REGION Network 297: CARRIER POWER UNIT DC LINK UNDERVOLTAGE
   RUNG wire#powerrail
      { S7_Templates := "SrcType := Word" } EQ_Contact(in1 := "DB101_DB_SDC_FAULTS".Carrier_Fault[8], in2 := 182)
      Coil( "DB302_HMI_Faults".Carrier8_Faults_1.%X11 )
   END_RUNG
   // the same network as SCL:
   "DB302_HMI_Faults".Carrier8_Faults_1.%X11 := "DB101_DB_SDC_FAULTS".Carrier_Fault[8] = 182;
END_REGION

REGION Network 298: CARRIER POWER UNIT LINE PHASE FAILURE
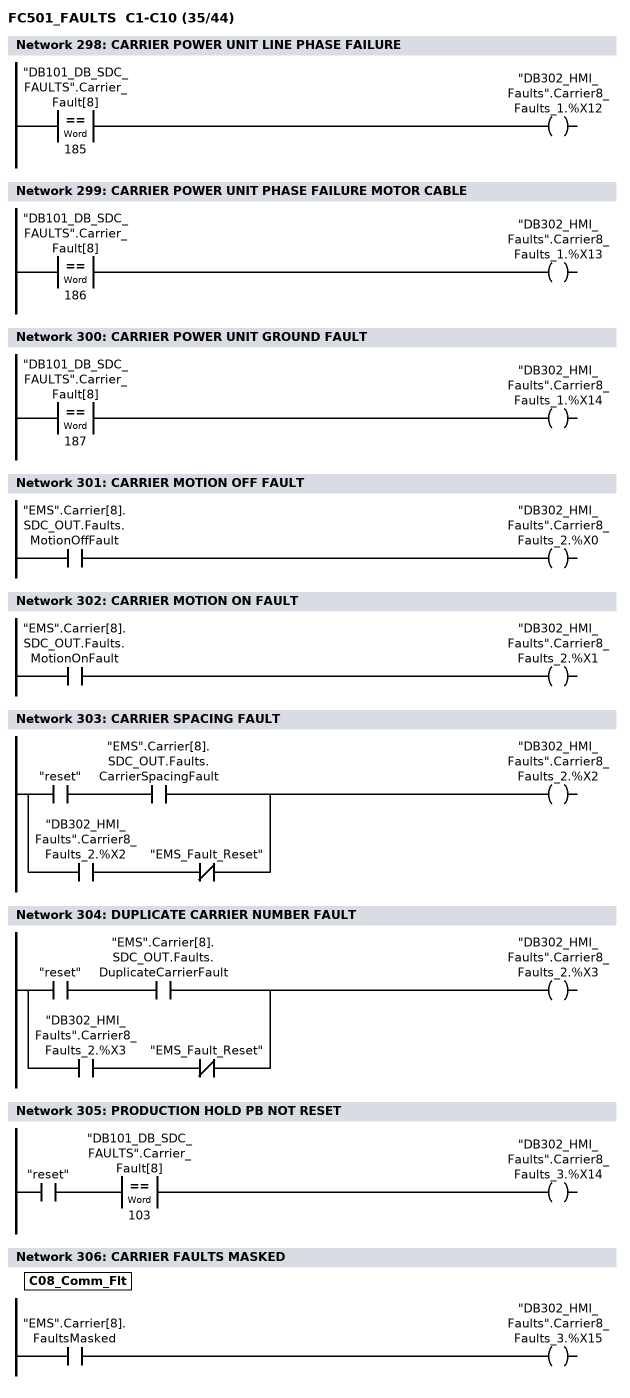
   RUNG wire#powerrail
      { S7_Templates := "SrcType := Word" } EQ_Contact(in1 := "DB101_DB_SDC_FAULTS".Carrier_Fault[8], in2 := 185)
      Coil( "DB302_HMI_Faults".Carrier8_Faults_1.%X12 )
   END_RUNG
   // the same network as SCL:
   "DB302_HMI_Faults".Carrier8_Faults_1.%X12 := "DB101_DB_SDC_FAULTS".Carrier_Fault[8] = 185;
END_REGION

REGION Network 299: CARRIER POWER UNIT PHASE FAILURE MOTOR CABLE
   RUNG wire#powerrail
      { S7_Templates := "SrcType := Word" } EQ_Contact(in1 := "DB101_DB_SDC_FAULTS".Carrier_Fault[8], in2 := 186)
      Coil( "DB302_HMI_Faults".Carrier8_Faults_1.%X13 )
   END_RUNG
   // the same network as SCL:
   "DB302_HMI_Faults".Carrier8_Faults_1.%X13 := "DB101_DB_SDC_FAULTS".Carrier_Fault[8] = 186;
END_REGION

REGION Network 300: CARRIER POWER UNIT GROUND FAULT
   RUNG wire#powerrail
      { S7_Templates := "SrcType := Word" } EQ_Contact(in1 := "DB101_DB_SDC_FAULTS".Carrier_Fault[8], in2 := 187)
      Coil( "DB302_HMI_Faults".Carrier8_Faults_1.%X14 )
   END_RUNG
   // the same network as SCL:
   "DB302_HMI_Faults".Carrier8_Faults_1.%X14 := "DB101_DB_SDC_FAULTS".Carrier_Fault[8] = 187;
END_REGION

REGION Network 301: CARRIER MOTION OFF FAULT
   RUNG wire#powerrail
      Contact( "EMS".Carrier[8].SDC_OUT.Faults.MotionOffFault )
      Coil( "DB302_HMI_Faults".Carrier8_Faults_2.%X0 )
   END_RUNG
   // the same network as SCL:
   "DB302_HMI_Faults".Carrier8_Faults_2.%X0 := "EMS".Carrier[8].SDC_OUT.Faults.MotionOffFault;
END_REGION

REGION Network 302: CARRIER MOTION ON FAULT
   RUNG wire#powerrail
      Contact( "EMS".Carrier[8].SDC_OUT.Faults.MotionOnFault )
      Coil( "DB302_HMI_Faults".Carrier8_Faults_2.%X1 )
   END_RUNG
   // the same network as SCL:
   "DB302_HMI_Faults".Carrier8_Faults_2.%X1 := "EMS".Carrier[8].SDC_OUT.Faults.MotionOnFault;
END_REGION

REGION Network 303: CARRIER SPACING FAULT
   RUNG wire#powerrail
      Contact( "reset" )
      Contact( "EMS".Carrier[8].SDC_OUT.Faults.CarrierSpacingFault )
      wire#w1
      Coil( "DB302_HMI_Faults".Carrier8_Faults_2.%X2 )
   END_RUNG
   RUNG wire#powerrail
      Contact( "DB302_HMI_Faults".Carrier8_Faults_2.%X2 )
      I_Contact( "EMS_Fault_Reset" )
   END_RUNG wire#w1
   // the same network as SCL:
   "DB302_HMI_Faults".Carrier8_Faults_2.%X2 := ("reset" AND "EMS".Carrier[8].SDC_OUT.Faults.CarrierSpacingFault) OR ("DB302_HMI_Faults".Carrier8_Faults_2.%X2 AND NOT "EMS_Fault_Reset");
END_REGION

REGION Network 304: DUPLICATE CARRIER NUMBER FAULT
   RUNG wire#powerrail
      Contact( "reset" )
      Contact( "EMS".Carrier[8].SDC_OUT.Faults.DuplicateCarrierFault )
      wire#w1
      Coil( "DB302_HMI_Faults".Carrier8_Faults_2.%X3 )
   END_RUNG
   RUNG wire#powerrail
      Contact( "DB302_HMI_Faults".Carrier8_Faults_2.%X3 )
      I_Contact( "EMS_Fault_Reset" )
   END_RUNG wire#w1
   // the same network as SCL:
   "DB302_HMI_Faults".Carrier8_Faults_2.%X3 := ("reset" AND "EMS".Carrier[8].SDC_OUT.Faults.DuplicateCarrierFault) OR ("DB302_HMI_Faults".Carrier8_Faults_2.%X3 AND NOT "EMS_Fault_Reset");
END_REGION

REGION Network 305: PRODUCTION HOLD PB NOT RESET
   RUNG wire#powerrail
      Contact( "reset" )
      { S7_Templates := "SrcType := Word" } EQ_Contact(in1 := "DB101_DB_SDC_FAULTS".Carrier_Fault[8], in2 := 103)
      Coil( "DB302_HMI_Faults".Carrier8_Faults_3.%X14 )
   END_RUNG
   // the same network as SCL:
   "DB302_HMI_Faults".Carrier8_Faults_3.%X14 := "reset" AND ("DB101_DB_SDC_FAULTS".Carrier_Fault[8] = 103);
END_REGION

REGION Network 306: CARRIER FAULTS MASKED
   Label( C08_Comm_Flt )
   RUNG wire#powerrail
      Contact( "EMS".Carrier[8].FaultsMasked )
      Coil( "DB302_HMI_Faults".Carrier8_Faults_3.%X15 )
   END_RUNG
   // the same network as SCL:
   C08_Comm_Flt:
   "DB302_HMI_Faults".Carrier8_Faults_3.%X15 := "EMS".Carrier[8].FaultsMasked;
END_REGION

REGION Network 307: CARRIER 9 FAULTS
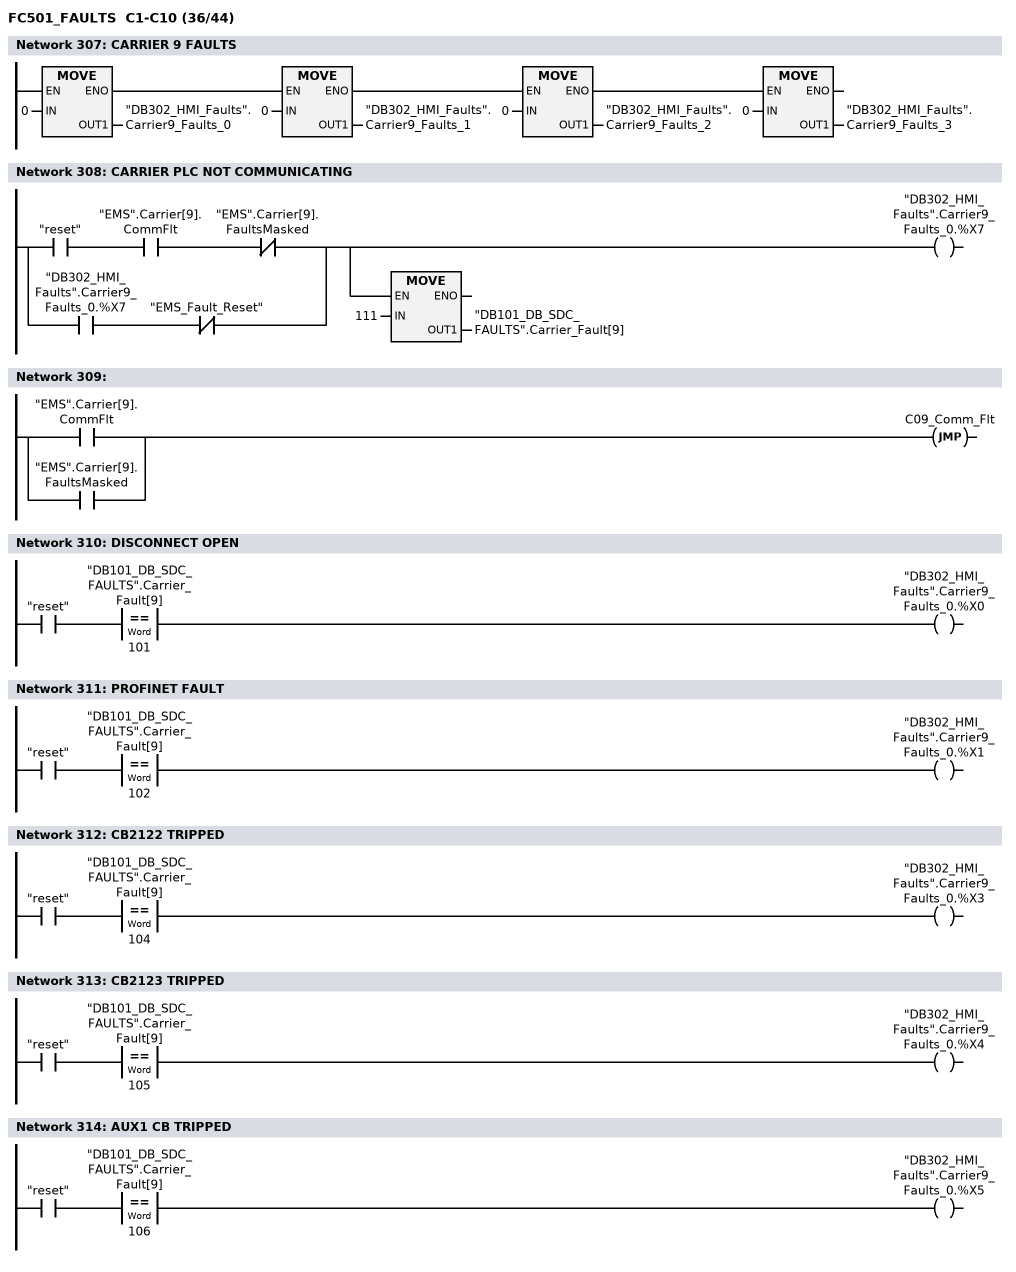
   RUNG wire#powerrail
      Move(in := 0, out1 => "DB302_HMI_Faults".Carrier9_Faults_0)
      Move(in := 0, out1 => "DB302_HMI_Faults".Carrier9_Faults_1)
      Move(in := 0, out1 => "DB302_HMI_Faults".Carrier9_Faults_2)
      Move(in := 0, out1 => "DB302_HMI_Faults".Carrier9_Faults_3)
   END_RUNG
   // the same network as SCL:
   "DB302_HMI_Faults".Carrier9_Faults_0 := 0;
   "DB302_HMI_Faults".Carrier9_Faults_1 := 0;
   "DB302_HMI_Faults".Carrier9_Faults_2 := 0;
   "DB302_HMI_Faults".Carrier9_Faults_3 := 0;
END_REGION

REGION Network 308: CARRIER PLC NOT COMMUNICATING
   RUNG wire#powerrail
      Contact( "reset" )
      Contact( "EMS".Carrier[9].CommFlt )
      I_Contact( "EMS".Carrier[9].FaultsMasked )
      wire#w1
      Coil( "DB302_HMI_Faults".Carrier9_Faults_0.%X7 )
   END_RUNG
   RUNG wire#powerrail
      Contact( "DB302_HMI_Faults".Carrier9_Faults_0.%X7 )
      I_Contact( "EMS_Fault_Reset" )
   END_RUNG wire#w1
   RUNG wire#w1
      Move(in := 111, out1 => "DB101_DB_SDC_FAULTS".Carrier_Fault[9])
   END_RUNG
   // the same network as SCL:
   "DB302_HMI_Faults".Carrier9_Faults_0.%X7 := ("reset" AND "EMS".Carrier[9].CommFlt AND NOT "EMS".Carrier[9].FaultsMasked) OR ("DB302_HMI_Faults".Carrier9_Faults_0.%X7 AND NOT "EMS_Fault_Reset");
   IF "DB302_HMI_Faults".Carrier9_Faults_0.%X7 THEN "DB101_DB_SDC_FAULTS".Carrier_Fault[9] := 111; END_IF;
END_REGION

REGION Network 309
   RUNG wire#powerrail
      Contact( "EMS".Carrier[9].CommFlt )
      wire#w1
      JumpCoil( C09_Comm_Flt )
   END_RUNG
   RUNG wire#powerrail
      Contact( "EMS".Carrier[9].FaultsMasked )
   END_RUNG wire#w1
   // the same network as SCL:
   IF "EMS".Carrier[9].CommFlt OR "EMS".Carrier[9].FaultsMasked THEN GOTO C09_Comm_Flt; END_IF;
END_REGION

REGION Network 310: DISCONNECT OPEN
   RUNG wire#powerrail
      Contact( "reset" )
      { S7_Templates := "SrcType := Word" } EQ_Contact(in1 := "DB101_DB_SDC_FAULTS".Carrier_Fault[9], in2 := 101)
      Coil( "DB302_HMI_Faults".Carrier9_Faults_0.%X0 )
   END_RUNG
   // the same network as SCL:
   "DB302_HMI_Faults".Carrier9_Faults_0.%X0 := "reset" AND ("DB101_DB_SDC_FAULTS".Carrier_Fault[9] = 101);
END_REGION

REGION Network 311: PROFINET FAULT
   RUNG wire#powerrail
      Contact( "reset" )
      { S7_Templates := "SrcType := Word" } EQ_Contact(in1 := "DB101_DB_SDC_FAULTS".Carrier_Fault[9], in2 := 102)
      Coil( "DB302_HMI_Faults".Carrier9_Faults_0.%X1 )
   END_RUNG
   // the same network as SCL:
   "DB302_HMI_Faults".Carrier9_Faults_0.%X1 := "reset" AND ("DB101_DB_SDC_FAULTS".Carrier_Fault[9] = 102);
END_REGION

REGION Network 312: CB2122 TRIPPED
   RUNG wire#powerrail
      Contact( "reset" )
      { S7_Templates := "SrcType := Word" } EQ_Contact(in1 := "DB101_DB_SDC_FAULTS".Carrier_Fault[9], in2 := 104)
      Coil( "DB302_HMI_Faults".Carrier9_Faults_0.%X3 )
   END_RUNG
   // the same network as SCL:
   "DB302_HMI_Faults".Carrier9_Faults_0.%X3 := "reset" AND ("DB101_DB_SDC_FAULTS".Carrier_Fault[9] = 104);
END_REGION

REGION Network 313: CB2123 TRIPPED
   RUNG wire#powerrail
      Contact( "reset" )
      { S7_Templates := "SrcType := Word" } EQ_Contact(in1 := "DB101_DB_SDC_FAULTS".Carrier_Fault[9], in2 := 105)
      Coil( "DB302_HMI_Faults".Carrier9_Faults_0.%X4 )
   END_RUNG
   // the same network as SCL:
   "DB302_HMI_Faults".Carrier9_Faults_0.%X4 := "reset" AND ("DB101_DB_SDC_FAULTS".Carrier_Fault[9] = 105);
END_REGION

REGION Network 314: AUX1 CB TRIPPED
   RUNG wire#powerrail
      Contact( "reset" )
      { S7_Templates := "SrcType := Word" } EQ_Contact(in1 := "DB101_DB_SDC_FAULTS".Carrier_Fault[9], in2 := 106)
      Coil( "DB302_HMI_Faults".Carrier9_Faults_0.%X5 )
   END_RUNG
   // the same network as SCL:
   "DB302_HMI_Faults".Carrier9_Faults_0.%X5 := "reset" AND ("DB101_DB_SDC_FAULTS".Carrier_Fault[9] = 106);
END_REGION

REGION Network 315: AUX2 CB TRIPPED
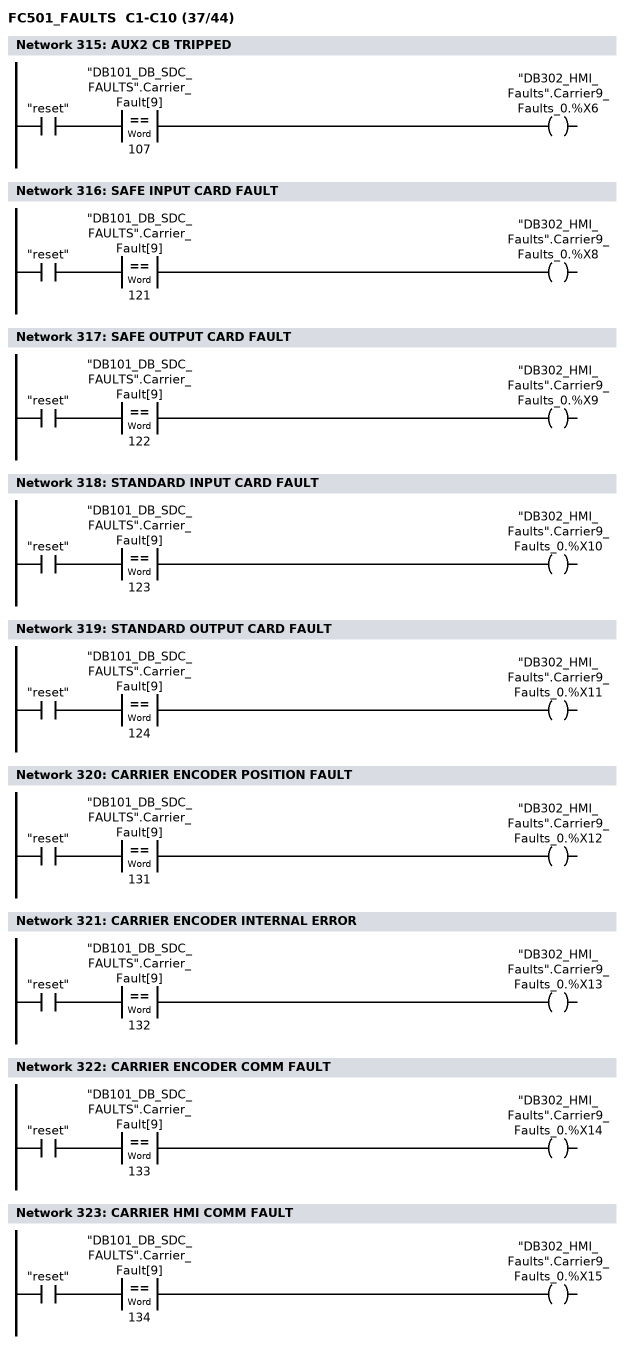
   RUNG wire#powerrail
      Contact( "reset" )
      { S7_Templates := "SrcType := Word" } EQ_Contact(in1 := "DB101_DB_SDC_FAULTS".Carrier_Fault[9], in2 := 107)
      Coil( "DB302_HMI_Faults".Carrier9_Faults_0.%X6 )
   END_RUNG
   // the same network as SCL:
   "DB302_HMI_Faults".Carrier9_Faults_0.%X6 := "reset" AND ("DB101_DB_SDC_FAULTS".Carrier_Fault[9] = 107);
END_REGION

REGION Network 316: SAFE INPUT CARD FAULT
   RUNG wire#powerrail
      Contact( "reset" )
      { S7_Templates := "SrcType := Word" } EQ_Contact(in1 := "DB101_DB_SDC_FAULTS".Carrier_Fault[9], in2 := 121)
      Coil( "DB302_HMI_Faults".Carrier9_Faults_0.%X8 )
   END_RUNG
   // the same network as SCL:
   "DB302_HMI_Faults".Carrier9_Faults_0.%X8 := "reset" AND ("DB101_DB_SDC_FAULTS".Carrier_Fault[9] = 121);
END_REGION

REGION Network 317: SAFE OUTPUT CARD FAULT
   RUNG wire#powerrail
      Contact( "reset" )
      { S7_Templates := "SrcType := Word" } EQ_Contact(in1 := "DB101_DB_SDC_FAULTS".Carrier_Fault[9], in2 := 122)
      Coil( "DB302_HMI_Faults".Carrier9_Faults_0.%X9 )
   END_RUNG
   // the same network as SCL:
   "DB302_HMI_Faults".Carrier9_Faults_0.%X9 := "reset" AND ("DB101_DB_SDC_FAULTS".Carrier_Fault[9] = 122);
END_REGION

REGION Network 318: STANDARD INPUT CARD FAULT
   RUNG wire#powerrail
      Contact( "reset" )
      { S7_Templates := "SrcType := Word" } EQ_Contact(in1 := "DB101_DB_SDC_FAULTS".Carrier_Fault[9], in2 := 123)
      Coil( "DB302_HMI_Faults".Carrier9_Faults_0.%X10 )
   END_RUNG
   // the same network as SCL:
   "DB302_HMI_Faults".Carrier9_Faults_0.%X10 := "reset" AND ("DB101_DB_SDC_FAULTS".Carrier_Fault[9] = 123);
END_REGION

REGION Network 319: STANDARD OUTPUT CARD FAULT
   RUNG wire#powerrail
      Contact( "reset" )
      { S7_Templates := "SrcType := Word" } EQ_Contact(in1 := "DB101_DB_SDC_FAULTS".Carrier_Fault[9], in2 := 124)
      Coil( "DB302_HMI_Faults".Carrier9_Faults_0.%X11 )
   END_RUNG
   // the same network as SCL:
   "DB302_HMI_Faults".Carrier9_Faults_0.%X11 := "reset" AND ("DB101_DB_SDC_FAULTS".Carrier_Fault[9] = 124);
END_REGION

REGION Network 320: CARRIER ENCODER POSITION FAULT
   RUNG wire#powerrail
      Contact( "reset" )
      { S7_Templates := "SrcType := Word" } EQ_Contact(in1 := "DB101_DB_SDC_FAULTS".Carrier_Fault[9], in2 := 131)
      Coil( "DB302_HMI_Faults".Carrier9_Faults_0.%X12 )
   END_RUNG
   // the same network as SCL:
   "DB302_HMI_Faults".Carrier9_Faults_0.%X12 := "reset" AND ("DB101_DB_SDC_FAULTS".Carrier_Fault[9] = 131);
END_REGION

REGION Network 321: CARRIER ENCODER INTERNAL ERROR
   RUNG wire#powerrail
      Contact( "reset" )
      { S7_Templates := "SrcType := Word" } EQ_Contact(in1 := "DB101_DB_SDC_FAULTS".Carrier_Fault[9], in2 := 132)
      Coil( "DB302_HMI_Faults".Carrier9_Faults_0.%X13 )
   END_RUNG
   // the same network as SCL:
   "DB302_HMI_Faults".Carrier9_Faults_0.%X13 := "reset" AND ("DB101_DB_SDC_FAULTS".Carrier_Fault[9] = 132);
END_REGION

REGION Network 322: CARRIER ENCODER COMM FAULT
   RUNG wire#powerrail
      Contact( "reset" )
      { S7_Templates := "SrcType := Word" } EQ_Contact(in1 := "DB101_DB_SDC_FAULTS".Carrier_Fault[9], in2 := 133)
      Coil( "DB302_HMI_Faults".Carrier9_Faults_0.%X14 )
   END_RUNG
   // the same network as SCL:
   "DB302_HMI_Faults".Carrier9_Faults_0.%X14 := "reset" AND ("DB101_DB_SDC_FAULTS".Carrier_Fault[9] = 133);
END_REGION

REGION Network 323: CARRIER HMI COMM FAULT
   RUNG wire#powerrail
      Contact( "reset" )
      { S7_Templates := "SrcType := Word" } EQ_Contact(in1 := "DB101_DB_SDC_FAULTS".Carrier_Fault[9], in2 := 134)
      Coil( "DB302_HMI_Faults".Carrier9_Faults_0.%X15 )
   END_RUNG
   // the same network as SCL:
   "DB302_HMI_Faults".Carrier9_Faults_0.%X15 := "reset" AND ("DB101_DB_SDC_FAULTS".Carrier_Fault[9] = 134);
END_REGION

REGION Network 324: CARRIER CRASH DETECTION FAULT
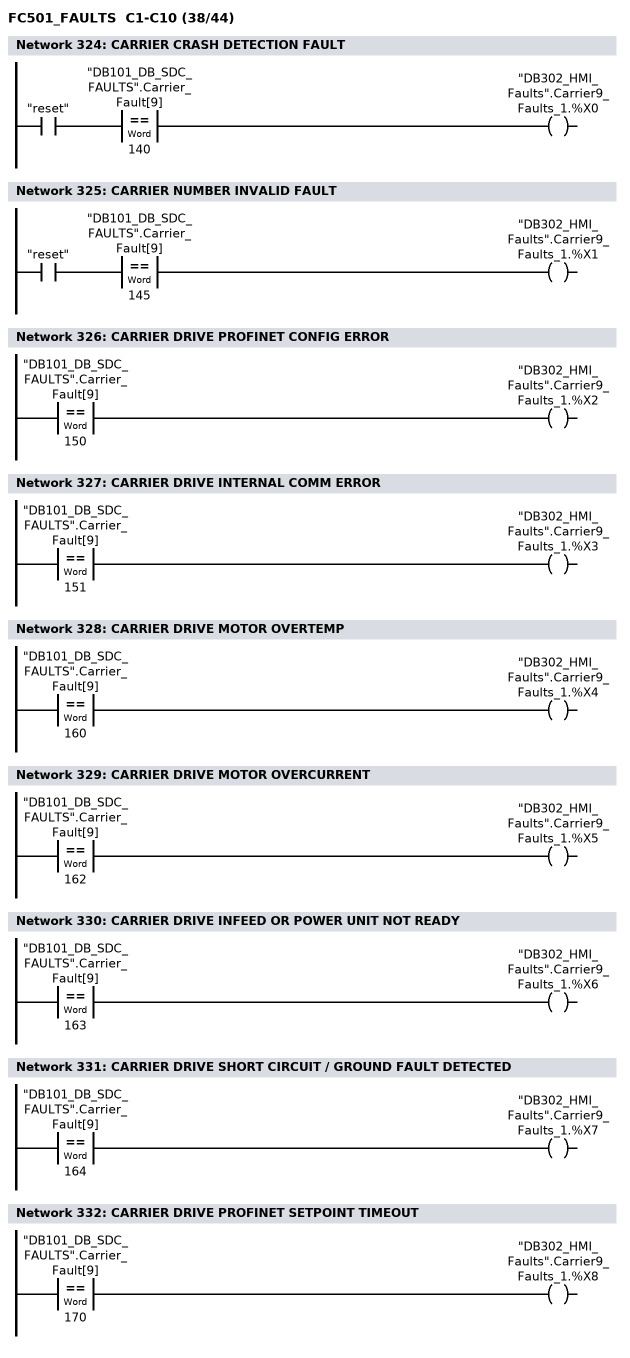
   RUNG wire#powerrail
      Contact( "reset" )
      { S7_Templates := "SrcType := Word" } EQ_Contact(in1 := "DB101_DB_SDC_FAULTS".Carrier_Fault[9], in2 := 140)
      Coil( "DB302_HMI_Faults".Carrier9_Faults_1.%X0 )
   END_RUNG
   // the same network as SCL:
   "DB302_HMI_Faults".Carrier9_Faults_1.%X0 := "reset" AND ("DB101_DB_SDC_FAULTS".Carrier_Fault[9] = 140);
END_REGION

REGION Network 325: CARRIER NUMBER INVALID FAULT
   RUNG wire#powerrail
      Contact( "reset" )
      { S7_Templates := "SrcType := Word" } EQ_Contact(in1 := "DB101_DB_SDC_FAULTS".Carrier_Fault[9], in2 := 145)
      Coil( "DB302_HMI_Faults".Carrier9_Faults_1.%X1 )
   END_RUNG
   // the same network as SCL:
   "DB302_HMI_Faults".Carrier9_Faults_1.%X1 := "reset" AND ("DB101_DB_SDC_FAULTS".Carrier_Fault[9] = 145);
END_REGION

REGION Network 326: CARRIER DRIVE PROFINET CONFIG ERROR
   RUNG wire#powerrail
      { S7_Templates := "SrcType := Word" } EQ_Contact(in1 := "DB101_DB_SDC_FAULTS".Carrier_Fault[9], in2 := 150)
      Coil( "DB302_HMI_Faults".Carrier9_Faults_1.%X2 )
   END_RUNG
   // the same network as SCL:
   "DB302_HMI_Faults".Carrier9_Faults_1.%X2 := "DB101_DB_SDC_FAULTS".Carrier_Fault[9] = 150;
END_REGION

REGION Network 327: CARRIER DRIVE INTERNAL COMM ERROR
   RUNG wire#powerrail
      { S7_Templates := "SrcType := Word" } EQ_Contact(in1 := "DB101_DB_SDC_FAULTS".Carrier_Fault[9], in2 := 151)
      Coil( "DB302_HMI_Faults".Carrier9_Faults_1.%X3 )
   END_RUNG
   // the same network as SCL:
   "DB302_HMI_Faults".Carrier9_Faults_1.%X3 := "DB101_DB_SDC_FAULTS".Carrier_Fault[9] = 151;
END_REGION

REGION Network 328: CARRIER DRIVE MOTOR OVERTEMP
   RUNG wire#powerrail
      { S7_Templates := "SrcType := Word" } EQ_Contact(in1 := "DB101_DB_SDC_FAULTS".Carrier_Fault[9], in2 := 160)
      Coil( "DB302_HMI_Faults".Carrier9_Faults_1.%X4 )
   END_RUNG
   // the same network as SCL:
   "DB302_HMI_Faults".Carrier9_Faults_1.%X4 := "DB101_DB_SDC_FAULTS".Carrier_Fault[9] = 160;
END_REGION

REGION Network 329: CARRIER DRIVE MOTOR OVERCURRENT
   RUNG wire#powerrail
      { S7_Templates := "SrcType := Word" } EQ_Contact(in1 := "DB101_DB_SDC_FAULTS".Carrier_Fault[9], in2 := 162)
      Coil( "DB302_HMI_Faults".Carrier9_Faults_1.%X5 )
   END_RUNG
   // the same network as SCL:
   "DB302_HMI_Faults".Carrier9_Faults_1.%X5 := "DB101_DB_SDC_FAULTS".Carrier_Fault[9] = 162;
END_REGION

REGION Network 330: CARRIER DRIVE INFEED OR POWER UNIT NOT READY
   RUNG wire#powerrail
      { S7_Templates := "SrcType := Word" } EQ_Contact(in1 := "DB101_DB_SDC_FAULTS".Carrier_Fault[9], in2 := 163)
      Coil( "DB302_HMI_Faults".Carrier9_Faults_1.%X6 )
   END_RUNG
   // the same network as SCL:
   "DB302_HMI_Faults".Carrier9_Faults_1.%X6 := "DB101_DB_SDC_FAULTS".Carrier_Fault[9] = 163;
END_REGION

REGION Network 331: CARRIER DRIVE SHORT CIRCUIT / GROUND FAULT DETECTED
   RUNG wire#powerrail
      { S7_Templates := "SrcType := Word" } EQ_Contact(in1 := "DB101_DB_SDC_FAULTS".Carrier_Fault[9], in2 := 164)
      Coil( "DB302_HMI_Faults".Carrier9_Faults_1.%X7 )
   END_RUNG
   // the same network as SCL:
   "DB302_HMI_Faults".Carrier9_Faults_1.%X7 := "DB101_DB_SDC_FAULTS".Carrier_Fault[9] = 164;
END_REGION

REGION Network 332: CARRIER DRIVE PROFINET SETPOINT TIMEOUT
   RUNG wire#powerrail
      { S7_Templates := "SrcType := Word" } EQ_Contact(in1 := "DB101_DB_SDC_FAULTS".Carrier_Fault[9], in2 := 170)
      Coil( "DB302_HMI_Faults".Carrier9_Faults_1.%X8 )
   END_RUNG
   // the same network as SCL:
   "DB302_HMI_Faults".Carrier9_Faults_1.%X8 := "DB101_DB_SDC_FAULTS".Carrier_Fault[9] = 170;
END_REGION

REGION Network 333: CARRIER POWER UNIT OVERCURRENT
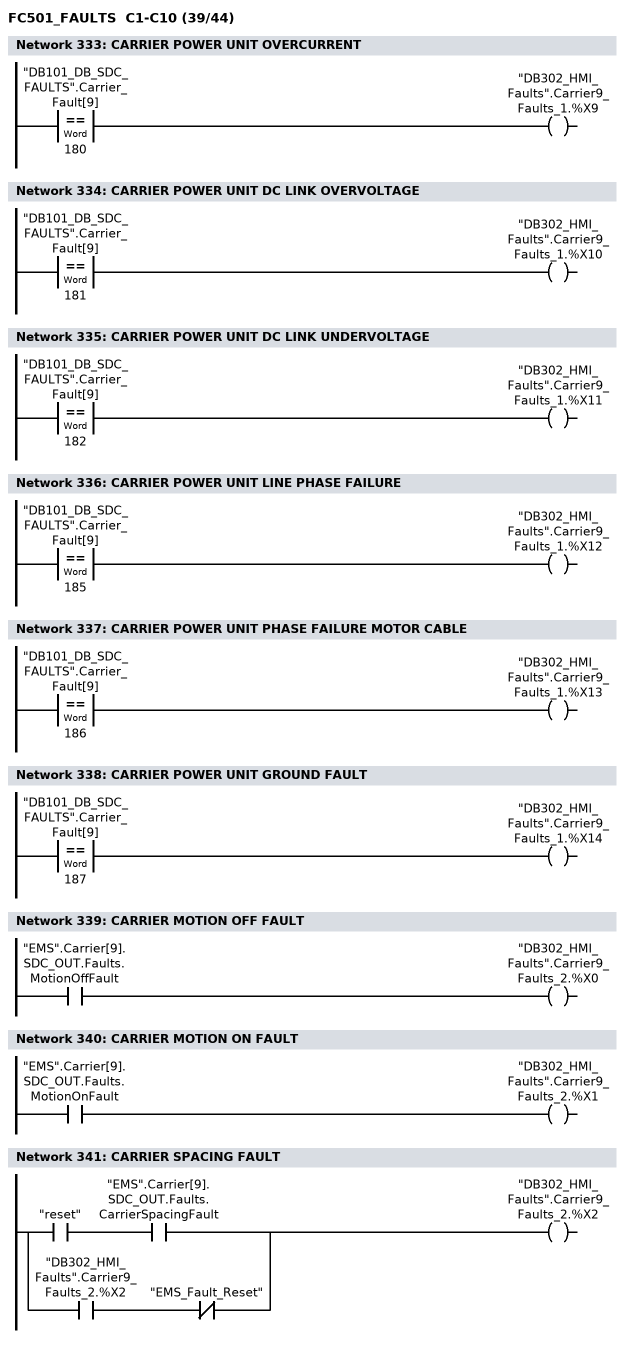
   RUNG wire#powerrail
      { S7_Templates := "SrcType := Word" } EQ_Contact(in1 := "DB101_DB_SDC_FAULTS".Carrier_Fault[9], in2 := 180)
      Coil( "DB302_HMI_Faults".Carrier9_Faults_1.%X9 )
   END_RUNG
   // the same network as SCL:
   "DB302_HMI_Faults".Carrier9_Faults_1.%X9 := "DB101_DB_SDC_FAULTS".Carrier_Fault[9] = 180;
END_REGION

REGION Network 334: CARRIER POWER UNIT DC LINK OVERVOLTAGE
   RUNG wire#powerrail
      { S7_Templates := "SrcType := Word" } EQ_Contact(in1 := "DB101_DB_SDC_FAULTS".Carrier_Fault[9], in2 := 181)
      Coil( "DB302_HMI_Faults".Carrier9_Faults_1.%X10 )
   END_RUNG
   // the same network as SCL:
   "DB302_HMI_Faults".Carrier9_Faults_1.%X10 := "DB101_DB_SDC_FAULTS".Carrier_Fault[9] = 181;
END_REGION

REGION Network 335: CARRIER POWER UNIT DC LINK UNDERVOLTAGE
   RUNG wire#powerrail
      { S7_Templates := "SrcType := Word" } EQ_Contact(in1 := "DB101_DB_SDC_FAULTS".Carrier_Fault[9], in2 := 182)
      Coil( "DB302_HMI_Faults".Carrier9_Faults_1.%X11 )
   END_RUNG
   // the same network as SCL:
   "DB302_HMI_Faults".Carrier9_Faults_1.%X11 := "DB101_DB_SDC_FAULTS".Carrier_Fault[9] = 182;
END_REGION

REGION Network 336: CARRIER POWER UNIT LINE PHASE FAILURE
   RUNG wire#powerrail
      { S7_Templates := "SrcType := Word" } EQ_Contact(in1 := "DB101_DB_SDC_FAULTS".Carrier_Fault[9], in2 := 185)
      Coil( "DB302_HMI_Faults".Carrier9_Faults_1.%X12 )
   END_RUNG
   // the same network as SCL:
   "DB302_HMI_Faults".Carrier9_Faults_1.%X12 := "DB101_DB_SDC_FAULTS".Carrier_Fault[9] = 185;
END_REGION

REGION Network 337: CARRIER POWER UNIT PHASE FAILURE MOTOR CABLE
   RUNG wire#powerrail
      { S7_Templates := "SrcType := Word" } EQ_Contact(in1 := "DB101_DB_SDC_FAULTS".Carrier_Fault[9], in2 := 186)
      Coil( "DB302_HMI_Faults".Carrier9_Faults_1.%X13 )
   END_RUNG
   // the same network as SCL:
   "DB302_HMI_Faults".Carrier9_Faults_1.%X13 := "DB101_DB_SDC_FAULTS".Carrier_Fault[9] = 186;
END_REGION

REGION Network 338: CARRIER POWER UNIT GROUND FAULT
   RUNG wire#powerrail
      { S7_Templates := "SrcType := Word" } EQ_Contact(in1 := "DB101_DB_SDC_FAULTS".Carrier_Fault[9], in2 := 187)
      Coil( "DB302_HMI_Faults".Carrier9_Faults_1.%X14 )
   END_RUNG
   // the same network as SCL:
   "DB302_HMI_Faults".Carrier9_Faults_1.%X14 := "DB101_DB_SDC_FAULTS".Carrier_Fault[9] = 187;
END_REGION

REGION Network 339: CARRIER MOTION OFF FAULT
   RUNG wire#powerrail
      Contact( "EMS".Carrier[9].SDC_OUT.Faults.MotionOffFault )
      Coil( "DB302_HMI_Faults".Carrier9_Faults_2.%X0 )
   END_RUNG
   // the same network as SCL:
   "DB302_HMI_Faults".Carrier9_Faults_2.%X0 := "EMS".Carrier[9].SDC_OUT.Faults.MotionOffFault;
END_REGION

REGION Network 340: CARRIER MOTION ON FAULT
   RUNG wire#powerrail
      Contact( "EMS".Carrier[9].SDC_OUT.Faults.MotionOnFault )
      Coil( "DB302_HMI_Faults".Carrier9_Faults_2.%X1 )
   END_RUNG
   // the same network as SCL:
   "DB302_HMI_Faults".Carrier9_Faults_2.%X1 := "EMS".Carrier[9].SDC_OUT.Faults.MotionOnFault;
END_REGION

REGION Network 341: CARRIER SPACING FAULT
   RUNG wire#powerrail
      Contact( "reset" )
      Contact( "EMS".Carrier[9].SDC_OUT.Faults.CarrierSpacingFault )
      wire#w1
      Coil( "DB302_HMI_Faults".Carrier9_Faults_2.%X2 )
   END_RUNG
   RUNG wire#powerrail
      Contact( "DB302_HMI_Faults".Carrier9_Faults_2.%X2 )
      I_Contact( "EMS_Fault_Reset" )
   END_RUNG wire#w1
   // the same network as SCL:
   "DB302_HMI_Faults".Carrier9_Faults_2.%X2 := ("reset" AND "EMS".Carrier[9].SDC_OUT.Faults.CarrierSpacingFault) OR ("DB302_HMI_Faults".Carrier9_Faults_2.%X2 AND NOT "EMS_Fault_Reset");
END_REGION

REGION Network 342: DUPLICATE CARRIER NUMBER FAULT
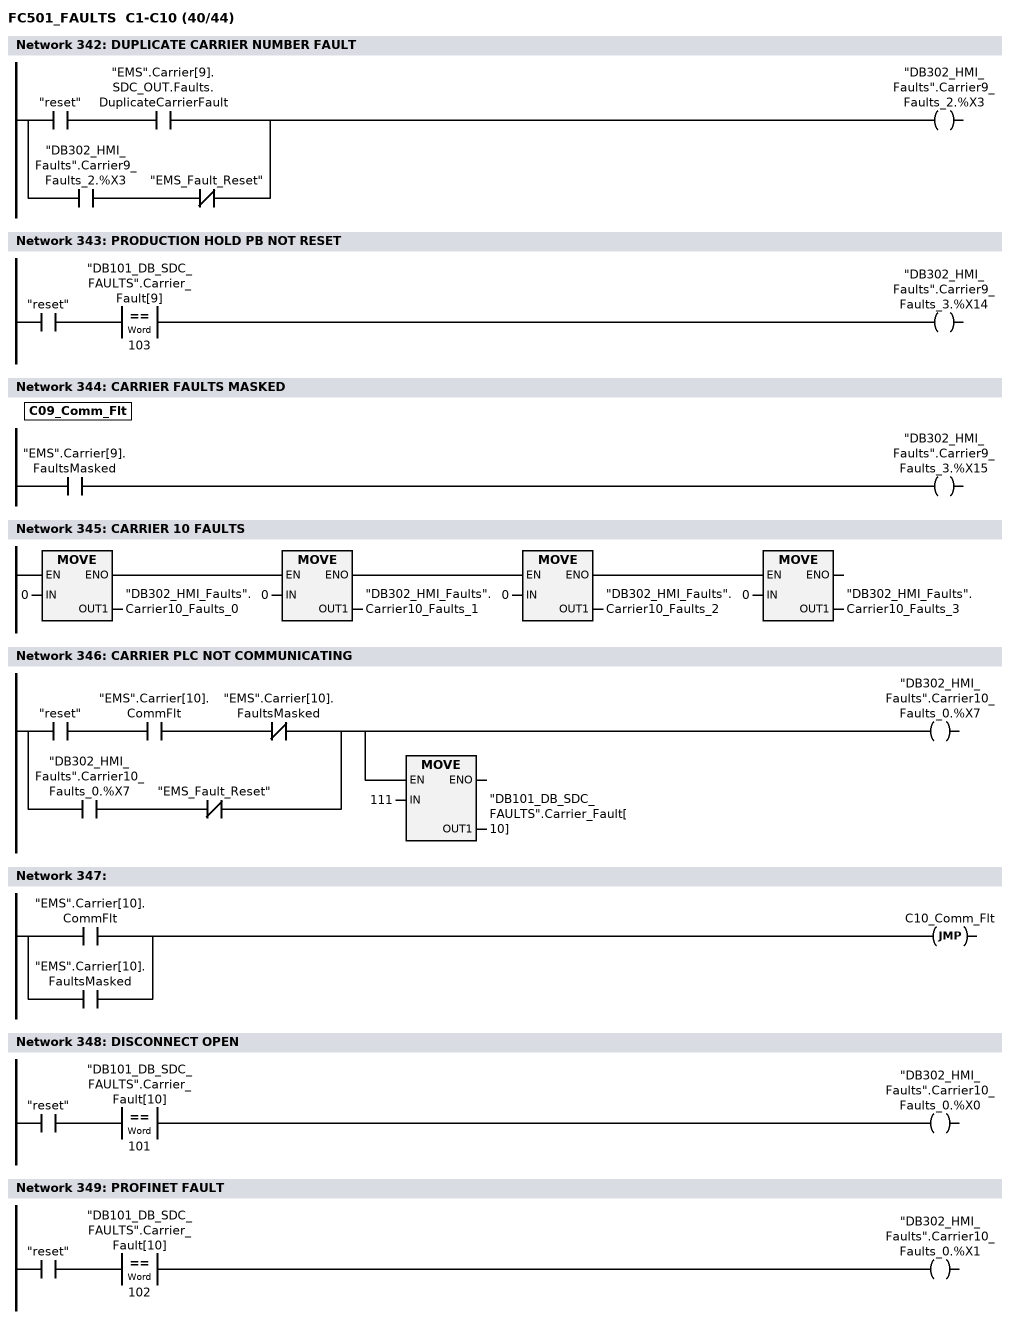
   RUNG wire#powerrail
      Contact( "reset" )
      Contact( "EMS".Carrier[9].SDC_OUT.Faults.DuplicateCarrierFault )
      wire#w1
      Coil( "DB302_HMI_Faults".Carrier9_Faults_2.%X3 )
   END_RUNG
   RUNG wire#powerrail
      Contact( "DB302_HMI_Faults".Carrier9_Faults_2.%X3 )
      I_Contact( "EMS_Fault_Reset" )
   END_RUNG wire#w1
   // the same network as SCL:
   "DB302_HMI_Faults".Carrier9_Faults_2.%X3 := ("reset" AND "EMS".Carrier[9].SDC_OUT.Faults.DuplicateCarrierFault) OR ("DB302_HMI_Faults".Carrier9_Faults_2.%X3 AND NOT "EMS_Fault_Reset");
END_REGION

REGION Network 343: PRODUCTION HOLD PB NOT RESET
   RUNG wire#powerrail
      Contact( "reset" )
      { S7_Templates := "SrcType := Word" } EQ_Contact(in1 := "DB101_DB_SDC_FAULTS".Carrier_Fault[9], in2 := 103)
      Coil( "DB302_HMI_Faults".Carrier9_Faults_3.%X14 )
   END_RUNG
   // the same network as SCL:
   "DB302_HMI_Faults".Carrier9_Faults_3.%X14 := "reset" AND ("DB101_DB_SDC_FAULTS".Carrier_Fault[9] = 103);
END_REGION

REGION Network 344: CARRIER FAULTS MASKED
   Label( C09_Comm_Flt )
   RUNG wire#powerrail
      Contact( "EMS".Carrier[9].FaultsMasked )
      Coil( "DB302_HMI_Faults".Carrier9_Faults_3.%X15 )
   END_RUNG
   // the same network as SCL:
   C09_Comm_Flt:
   "DB302_HMI_Faults".Carrier9_Faults_3.%X15 := "EMS".Carrier[9].FaultsMasked;
END_REGION

REGION Network 345: CARRIER 10 FAULTS
   RUNG wire#powerrail
      Move(in := 0, out1 => "DB302_HMI_Faults".Carrier10_Faults_0)
      Move(in := 0, out1 => "DB302_HMI_Faults".Carrier10_Faults_1)
      Move(in := 0, out1 => "DB302_HMI_Faults".Carrier10_Faults_2)
      Move(in := 0, out1 => "DB302_HMI_Faults".Carrier10_Faults_3)
   END_RUNG
   // the same network as SCL:
   "DB302_HMI_Faults".Carrier10_Faults_0 := 0;
   "DB302_HMI_Faults".Carrier10_Faults_1 := 0;
   "DB302_HMI_Faults".Carrier10_Faults_2 := 0;
   "DB302_HMI_Faults".Carrier10_Faults_3 := 0;
END_REGION

REGION Network 346: CARRIER PLC NOT COMMUNICATING
   RUNG wire#powerrail
      Contact( "reset" )
      Contact( "EMS".Carrier[10].CommFlt )
      I_Contact( "EMS".Carrier[10].FaultsMasked )
      wire#w1
      Coil( "DB302_HMI_Faults".Carrier10_Faults_0.%X7 )
   END_RUNG
   RUNG wire#powerrail
      Contact( "DB302_HMI_Faults".Carrier10_Faults_0.%X7 )
      I_Contact( "EMS_Fault_Reset" )
   END_RUNG wire#w1
   RUNG wire#w1
      Move(in := 111, out1 => "DB101_DB_SDC_FAULTS".Carrier_Fault[10])
   END_RUNG
   // the same network as SCL:
   "DB302_HMI_Faults".Carrier10_Faults_0.%X7 := ("reset" AND "EMS".Carrier[10].CommFlt AND NOT "EMS".Carrier[10].FaultsMasked) OR ("DB302_HMI_Faults".Carrier10_Faults_0.%X7 AND NOT "EMS_Fault_Reset");
   IF "DB302_HMI_Faults".Carrier10_Faults_0.%X7 THEN "DB101_DB_SDC_FAULTS".Carrier_Fault[10] := 111; END_IF;
END_REGION

REGION Network 347
   RUNG wire#powerrail
      Contact( "EMS".Carrier[10].CommFlt )
      wire#w1
      JumpCoil( C10_Comm_Flt )
   END_RUNG
   RUNG wire#powerrail
      Contact( "EMS".Carrier[10].FaultsMasked )
   END_RUNG wire#w1
   // the same network as SCL:
   IF "EMS".Carrier[10].CommFlt OR "EMS".Carrier[10].FaultsMasked THEN GOTO C10_Comm_Flt; END_IF;
END_REGION

REGION Network 348: DISCONNECT OPEN
   RUNG wire#powerrail
      Contact( "reset" )
      { S7_Templates := "SrcType := Word" } EQ_Contact(in1 := "DB101_DB_SDC_FAULTS".Carrier_Fault[10], in2 := 101)
      Coil( "DB302_HMI_Faults".Carrier10_Faults_0.%X0 )
   END_RUNG
   // the same network as SCL:
   "DB302_HMI_Faults".Carrier10_Faults_0.%X0 := "reset" AND ("DB101_DB_SDC_FAULTS".Carrier_Fault[10] = 101);
END_REGION

REGION Network 349: PROFINET FAULT
   RUNG wire#powerrail
      Contact( "reset" )
      { S7_Templates := "SrcType := Word" } EQ_Contact(in1 := "DB101_DB_SDC_FAULTS".Carrier_Fault[10], in2 := 102)
      Coil( "DB302_HMI_Faults".Carrier10_Faults_0.%X1 )
   END_RUNG
   // the same network as SCL:
   "DB302_HMI_Faults".Carrier10_Faults_0.%X1 := "reset" AND ("DB101_DB_SDC_FAULTS".Carrier_Fault[10] = 102);
END_REGION

REGION Network 350: CB2122 TRIPPED
